   9: EQU(Seat_Auxiliary_Ch_Memory,-1)OTE(To_Sfty.Seat_Auxiliary_Ch_Memory);
END_ROUTINE

ROUTINE Main   (* ladder *)
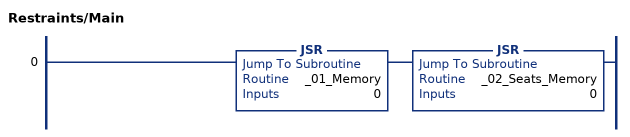
   0: JSR(_01_Memory,0)JSR(_02_Seats_Memory,0);
END_ROUTINE
END_PROGRAM

PROGRAM S_Alarms   (* main routine Main, safety *)
VAR
   LapBars_Alarms_Time : DINT := 2000;
   OS : DINT := 801;
   Timer : TIMER[60] := ([0].PRE := 2000, [1].PRE := 2000, [2].PRE := 2000, [3].PRE := 2000, [4].PRE := 2000, [5].PRE := 2000, [6].PRE := 2000, [7].PRE := 2000, [8].PRE := 2000, [8].ACC := 1520, [9].PRE := 5000, [10].PRE := 200, [11].PRE := 200, [12].PRE := 7000, [13].PRE := 5000, [14].PRE := 1000, [15].PRE := 20000, [16].PRE := 500, [17].PRE := 500, [18].PRE := 99999999, [19].PRE := 9000, [20].PRE := 2500, [21].PRE := 2500, [22].PRE := 5000, [23].PRE := 10000, [24].PRE := 5000, [25].PRE := 5000, [26].PRE := 100000, [27].PRE := 30000, [28].PRE := 2000, [29].PRE := 2000, [30].PRE := 2000, [31].PRE := 2000, [32].PRE := 2000, [33].PRE := 2000, [34].PRE := 2000, [35].PRE := 2000, [36].PRE := 2000, [37].PRE := 2000, [38].PRE := 60000, [39].PRE := 60000, [40].PRE := 7000, [41].PRE := 600, [42].PRE := 99999999, [43].PRE := 500, [44].PRE := 500, [45].PRE := 500);
        [18]   // Revolution time
        [16]   // Overspeed alarm pending activation from startup after direction change.
        [17]   // Overspeed alarm pending activation from startup after direction change.
        [19]   // Waiting for overspeed protection to be enabled at startup
        [43]   // Overspeed alarm pending activation from startup after direction change.
        [44]   // Overspeed alarm pending activation from startup after direction change.
   Timer_Restraints_Open : TIMER[41] := ([1].PRE := 200, [2].PRE := 200, [3].PRE := 200, [4].PRE := 200, [5].PRE := 200, [6].PRE := 200, [7].PRE := 200, [8].PRE := 200, [9].PRE := 200, [10].PRE := 200, [11].PRE := 200, [12].PRE := 200, [13].PRE := 200, [14].PRE := 200, [15].PRE := 200, [16].PRE := 200, [17].PRE := 200, [18].PRE := 200, [19].PRE := 200, [20].PRE := 200, [21].PRE := 200, [22].PRE := 200, [23].PRE := 200, [24].PRE := 200, [25].PRE := 200, [26].PRE := 200, [27].PRE := 200, [28].PRE := 200, [29].PRE := 200, [30].PRE := 200, [31].PRE := 200, [32].PRE := 200, [33].PRE := 200, [34].PRE := 200, [35].PRE := 200, [36].PRE := 200, [37].PRE := 200, [38].PRE := 200, [39].PRE := 200, [40].PRE := 200);
END_VAR

ROUTINE _00_Communication   (* ladder *)
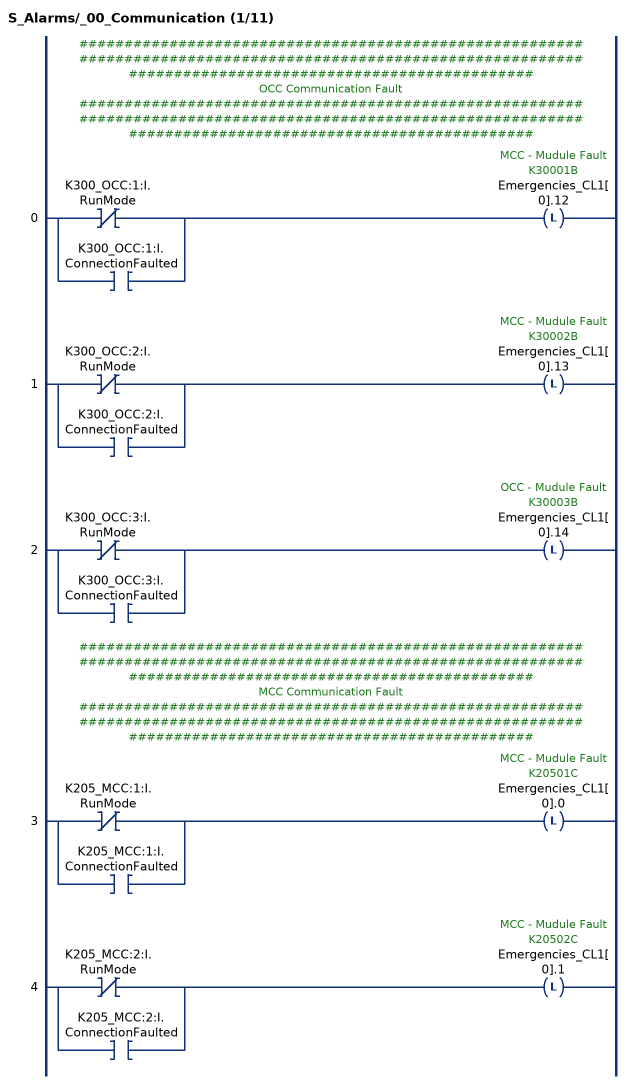
   // #############################################################################################################################################################
   // OCC Communication Fault
   // #############################################################################################################################################################
   0: [XIO(K300_OCC:1:I.RunMode) ,XIC(K300_OCC:1:I.ConnectionFaulted) ]OTL(Emergencies_CL1[0].12);
   1: [XIO(K300_OCC:2:I.RunMode) ,XIC(K300_OCC:2:I.ConnectionFaulted) ]OTL(Emergencies_CL1[0].13);
   2: [XIO(K300_OCC:3:I.RunMode) ,XIC(K300_OCC:3:I.ConnectionFaulted) ]OTL(Emergencies_CL1[0].14);
   // #############################################################################################################################################################
   // MCC Communication Fault
   // #############################################################################################################################################################
   3: [XIO(K205_MCC:1:I.RunMode) ,XIC(K205_MCC:1:I.ConnectionFaulted) ]OTL(Emergencies_CL1[0].0);
   4: [XIO(K205_MCC:2:I.RunMode) ,XIC(K205_MCC:2:I.ConnectionFaulted) ]OTL(Emergencies_CL1[0].1);
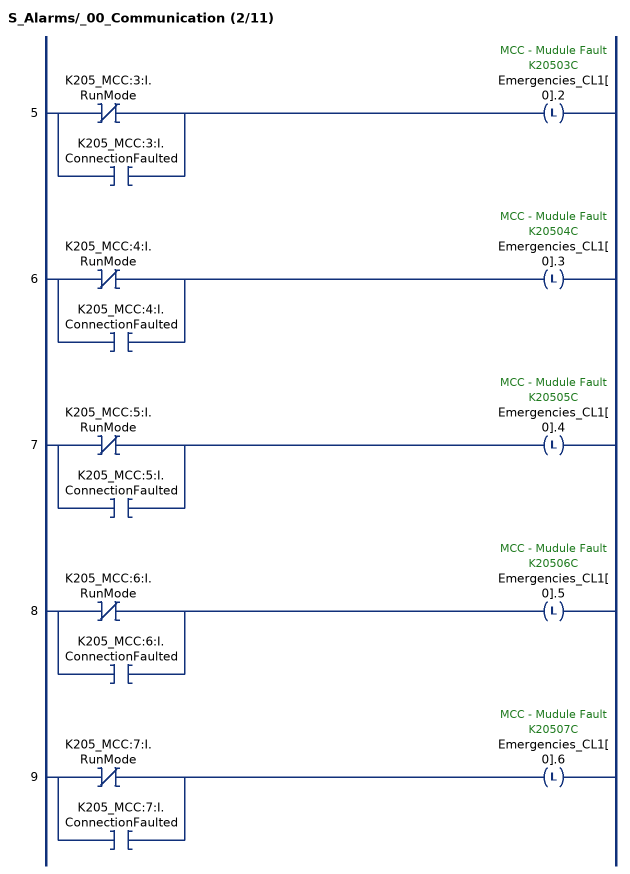
   5: [XIO(K205_MCC:3:I.RunMode) ,XIC(K205_MCC:3:I.ConnectionFaulted) ]OTL(Emergencies_CL1[0].2);
   6: [XIO(K205_MCC:4:I.RunMode) ,XIC(K205_MCC:4:I.ConnectionFaulted) ]OTL(Emergencies_CL1[0].3);
   7: [XIO(K205_MCC:5:I.RunMode) ,XIC(K205_MCC:5:I.ConnectionFaulted) ]OTL(Emergencies_CL1[0].4);
   8: [XIO(K205_MCC:6:I.RunMode) ,XIC(K205_MCC:6:I.ConnectionFaulted) ]OTL(Emergencies_CL1[0].5);
   9: [XIO(K205_MCC:7:I.RunMode) ,XIC(K205_MCC:7:I.ConnectionFaulted) ]OTL(Emergencies_CL1[0].6);
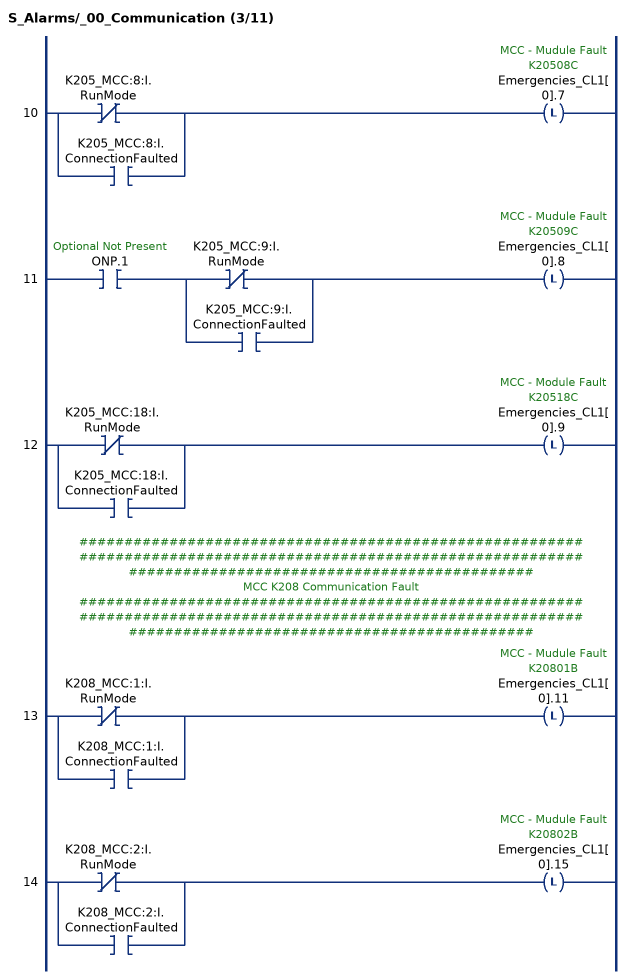
   10: [XIO(K205_MCC:8:I.RunMode) ,XIC(K205_MCC:8:I.ConnectionFaulted) ]OTL(Emergencies_CL1[0].7);
   11: XIC(ONP.1)[XIO(K205_MCC:9:I.RunMode) ,XIC(K205_MCC:9:I.ConnectionFaulted) ]OTL(Emergencies_CL1[0].8);
   12: [XIO(K205_MCC:18:I.RunMode) ,XIC(K205_MCC:18:I.ConnectionFaulted) ]OTL(Emergencies_CL1[0].9);
   // #############################################################################################################################################################
   // MCC K208 Communication Fault
   // #############################################################################################################################################################
   13: [XIO(K208_MCC:1:I.RunMode) ,XIC(K208_MCC:1:I.ConnectionFaulted) ]OTL(Emergencies_CL1[0].11);
   14: [XIO(K208_MCC:2:I.RunMode) ,XIC(K208_MCC:2:I.ConnectionFaulted) ]OTL(Emergencies_CL1[0].15);
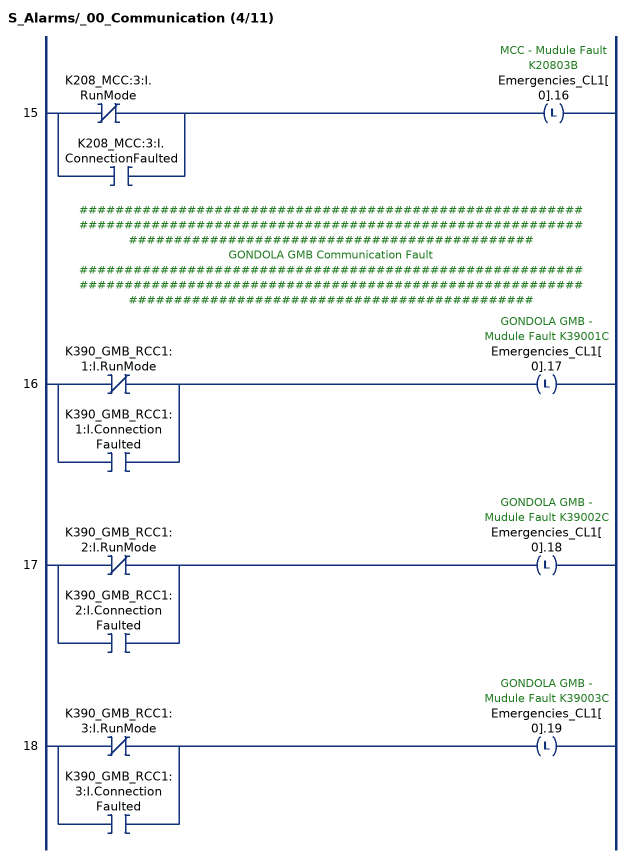
   15: [XIO(K208_MCC:3:I.RunMode) ,XIC(K208_MCC:3:I.ConnectionFaulted) ]OTL(Emergencies_CL1[0].16);
   // #############################################################################################################################################################
   // GONDOLA GMB Communication Fault
   // #############################################################################################################################################################
   16: [XIO(K390_GMB_RCC1:1:I.RunMode) ,XIC(K390_GMB_RCC1:1:I.ConnectionFaulted) ]OTL(Emergencies_CL1[0].17);
   17: [XIO(K390_GMB_RCC1:2:I.RunMode) ,XIC(K390_GMB_RCC1:2:I.ConnectionFaulted) ]OTL(Emergencies_CL1[0].18);
   18: [XIO(K390_GMB_RCC1:3:I.RunMode) ,XIC(K390_GMB_RCC1:3:I.ConnectionFaulted) ]OTL(Emergencies_CL1[0].19);
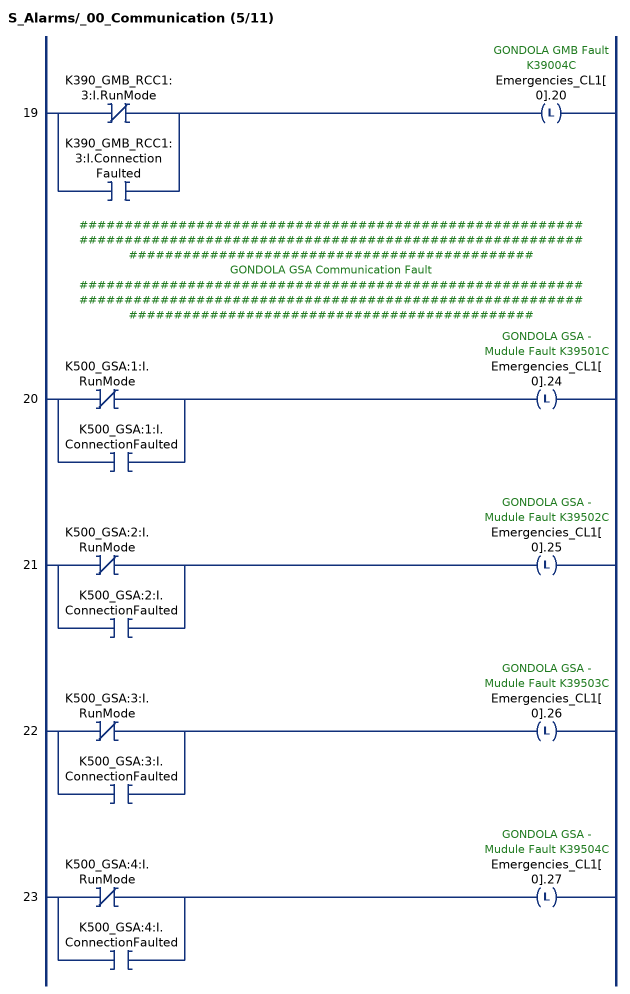
   19: [XIO(K390_GMB_RCC1:3:I.RunMode) ,XIC(K390_GMB_RCC1:3:I.ConnectionFaulted) ]OTL(Emergencies_CL1[0].20);
   // #############################################################################################################################################################
   // GONDOLA GSA Communication Fault
   // #############################################################################################################################################################
   20: [XIO(K500_GSA:1:I.RunMode) ,XIC(K500_GSA:1:I.ConnectionFaulted) ]OTL(Emergencies_CL1[0].24);
   21: [XIO(K500_GSA:2:I.RunMode) ,XIC(K500_GSA:2:I.ConnectionFaulted) ]OTL(Emergencies_CL1[0].25);
   22: [XIO(K500_GSA:3:I.RunMode) ,XIC(K500_GSA:3:I.ConnectionFaulted) ]OTL(Emergencies_CL1[0].26);
   23: [XIO(K500_GSA:4:I.RunMode) ,XIC(K500_GSA:4:I.ConnectionFaulted) ]OTL(Emergencies_CL1[0].27);
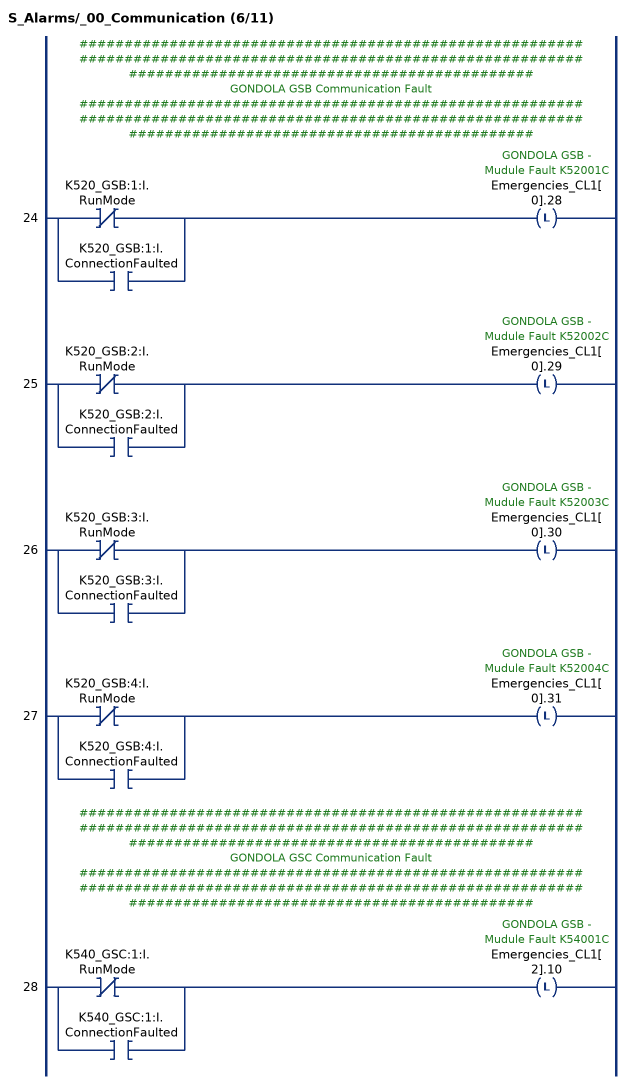
   // #############################################################################################################################################################
   // GONDOLA GSB Communication Fault
   // #############################################################################################################################################################
   24: [XIO(K520_GSB:1:I.RunMode) ,XIC(K520_GSB:1:I.ConnectionFaulted) ]OTL(Emergencies_CL1[0].28);
   25: [XIO(K520_GSB:2:I.RunMode) ,XIC(K520_GSB:2:I.ConnectionFaulted) ]OTL(Emergencies_CL1[0].29);
   26: [XIO(K520_GSB:3:I.RunMode) ,XIC(K520_GSB:3:I.ConnectionFaulted) ]OTL(Emergencies_CL1[0].30);
   27: [XIO(K520_GSB:4:I.RunMode) ,XIC(K520_GSB:4:I.ConnectionFaulted) ]OTL(Emergencies_CL1[0].31);
   // #############################################################################################################################################################
   // GONDOLA GSC Communication Fault
   // #############################################################################################################################################################
   28: [XIO(K540_GSC:1:I.RunMode) ,XIC(K540_GSC:1:I.ConnectionFaulted) ]OTL(Emergencies_CL1[2].10);
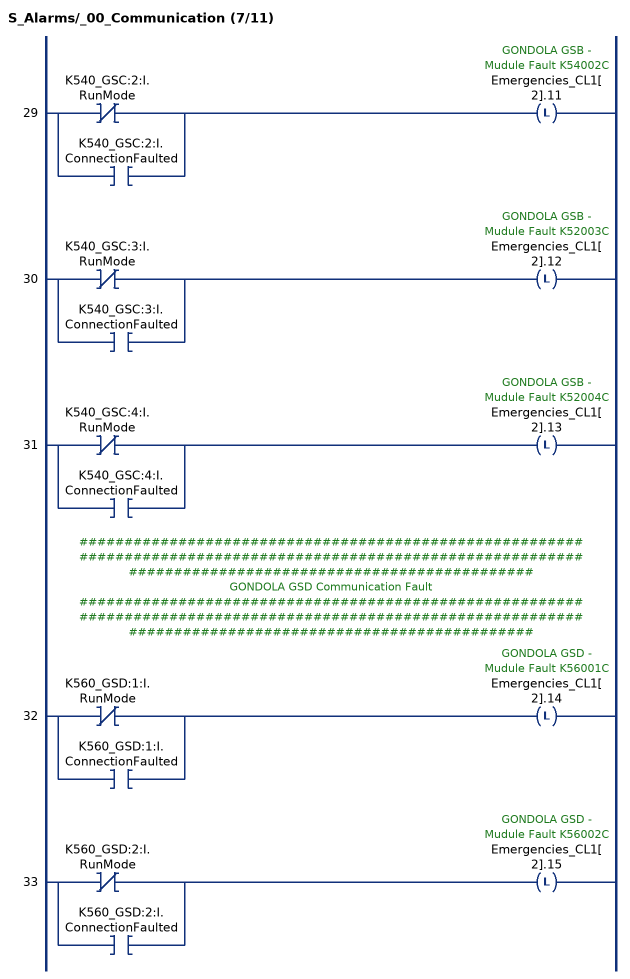
   29: [XIO(K540_GSC:2:I.RunMode) ,XIC(K540_GSC:2:I.ConnectionFaulted) ]OTL(Emergencies_CL1[2].11);
   30: [XIO(K540_GSC:3:I.RunMode) ,XIC(K540_GSC:3:I.ConnectionFaulted) ]OTL(Emergencies_CL1[2].12);
   31: [XIO(K540_GSC:4:I.RunMode) ,XIC(K540_GSC:4:I.ConnectionFaulted) ]OTL(Emergencies_CL1[2].13);
   // #############################################################################################################################################################
   // GONDOLA GSD Communication Fault
   // #############################################################################################################################################################
   32: [XIO(K560_GSD:1:I.RunMode) ,XIC(K560_GSD:1:I.ConnectionFaulted) ]OTL(Emergencies_CL1[2].14);
   33: [XIO(K560_GSD:2:I.RunMode) ,XIC(K560_GSD:2:I.ConnectionFaulted) ]OTL(Emergencies_CL1[2].15);
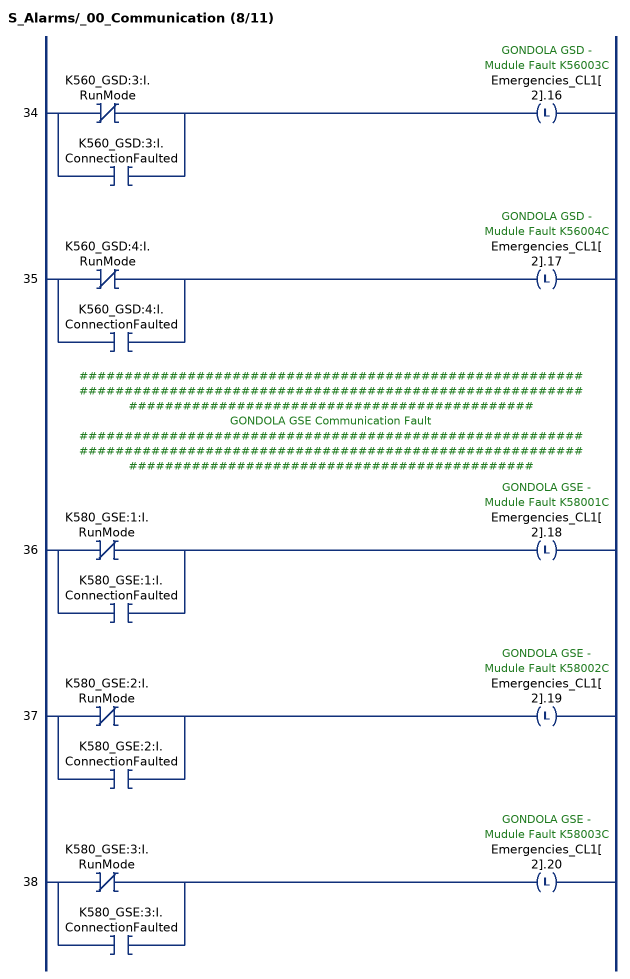
   34: [XIO(K560_GSD:3:I.RunMode) ,XIC(K560_GSD:3:I.ConnectionFaulted) ]OTL(Emergencies_CL1[2].16);
   35: [XIO(K560_GSD:4:I.RunMode) ,XIC(K560_GSD:4:I.ConnectionFaulted) ]OTL(Emergencies_CL1[2].17);
   // #############################################################################################################################################################
   // GONDOLA GSE Communication Fault
   // #############################################################################################################################################################
   36: [XIO(K580_GSE:1:I.RunMode) ,XIC(K580_GSE:1:I.ConnectionFaulted) ]OTL(Emergencies_CL1[2].18);
   37: [XIO(K580_GSE:2:I.RunMode) ,XIC(K580_GSE:2:I.ConnectionFaulted) ]OTL(Emergencies_CL1[2].19);
   38: [XIO(K580_GSE:3:I.RunMode) ,XIC(K580_GSE:3:I.ConnectionFaulted) ]OTL(Emergencies_CL1[2].20);
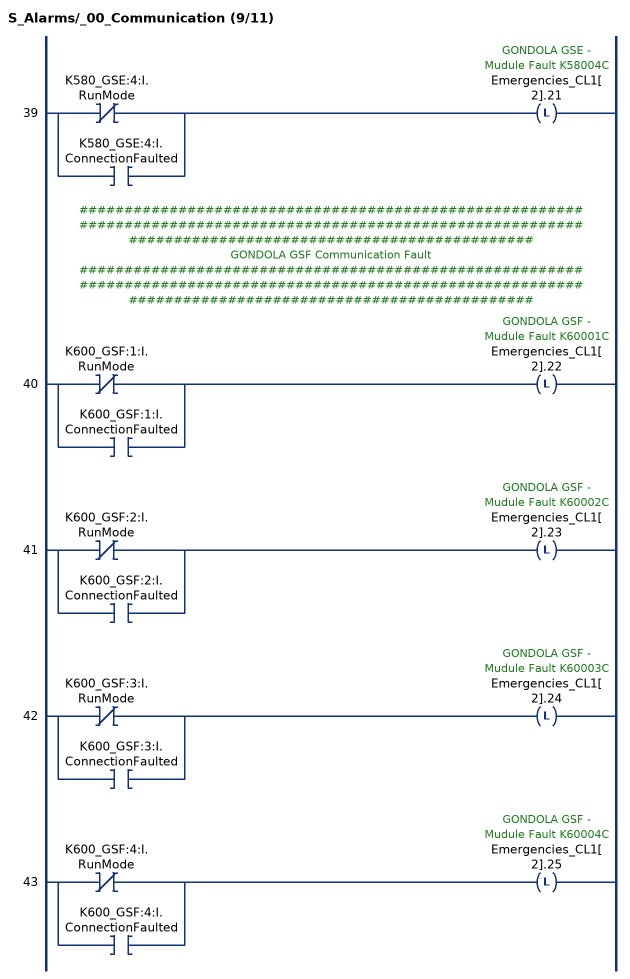
   39: [XIO(K580_GSE:4:I.RunMode) ,XIC(K580_GSE:4:I.ConnectionFaulted) ]OTL(Emergencies_CL1[2].21);
   // #############################################################################################################################################################
   // GONDOLA GSF Communication Fault
   // #############################################################################################################################################################
   40: [XIO(K600_GSF:1:I.RunMode) ,XIC(K600_GSF:1:I.ConnectionFaulted) ]OTL(Emergencies_CL1[2].22);
   41: [XIO(K600_GSF:2:I.RunMode) ,XIC(K600_GSF:2:I.ConnectionFaulted) ]OTL(Emergencies_CL1[2].23);
   42: [XIO(K600_GSF:3:I.RunMode) ,XIC(K600_GSF:3:I.ConnectionFaulted) ]OTL(Emergencies_CL1[2].24);
   43: [XIO(K600_GSF:4:I.RunMode) ,XIC(K600_GSF:4:I.ConnectionFaulted) ]OTL(Emergencies_CL1[2].25);
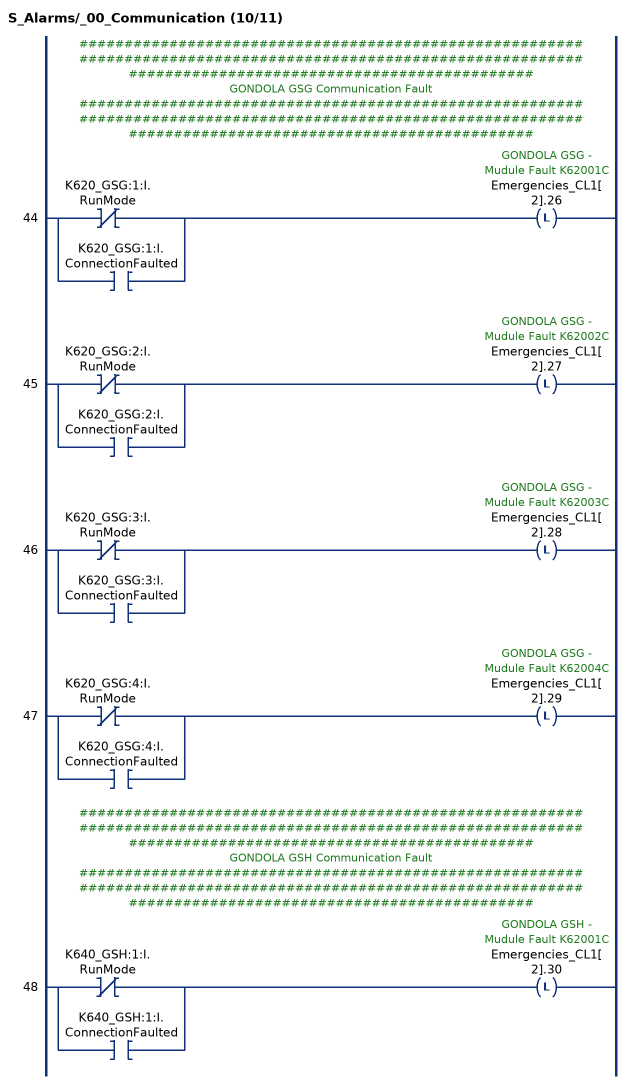
   // #############################################################################################################################################################
   // GONDOLA GSG Communication Fault
   // #############################################################################################################################################################
   44: [XIO(K620_GSG:1:I.RunMode) ,XIC(K620_GSG:1:I.ConnectionFaulted) ]OTL(Emergencies_CL1[2].26);
   45: [XIO(K620_GSG:2:I.RunMode) ,XIC(K620_GSG:2:I.ConnectionFaulted) ]OTL(Emergencies_CL1[2].27);
   46: [XIO(K620_GSG:3:I.RunMode) ,XIC(K620_GSG:3:I.ConnectionFaulted) ]OTL(Emergencies_CL1[2].28);
   47: [XIO(K620_GSG:4:I.RunMode) ,XIC(K620_GSG:4:I.ConnectionFaulted) ]OTL(Emergencies_CL1[2].29);
   // #############################################################################################################################################################
   // GONDOLA GSH Communication Fault
   // #############################################################################################################################################################
   48: [XIO(K640_GSH:1:I.RunMode) ,XIC(K640_GSH:1:I.ConnectionFaulted) ]OTL(Emergencies_CL1[2].30);
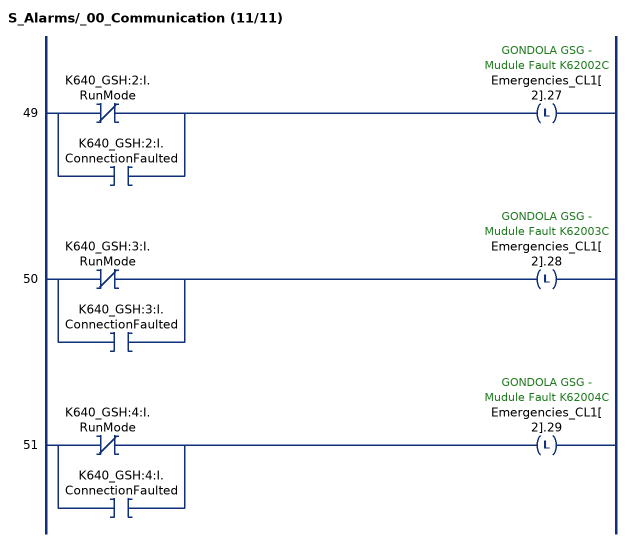
   49: [XIO(K640_GSH:2:I.RunMode) ,XIC(K640_GSH:2:I.ConnectionFaulted) ]OTL(Emergencies_CL1[2].27);
   50: [XIO(K640_GSH:3:I.RunMode) ,XIC(K640_GSH:3:I.ConnectionFaulted) ]OTL(Emergencies_CL1[2].28);
   51: [XIO(K640_GSH:4:I.RunMode) ,XIC(K640_GSH:4:I.ConnectionFaulted) ]OTL(Emergencies_CL1[2].29);
END_ROUTINE
